        [840] := 2776, [841] := 2780, [842] := 2778, [843] := 2773, [844] := 2778, [845] := 2776, [846] := 2780, [847] := 2783, [848] := 2766, [849] := 2787, [850] := 2773, [851] := 2776, [852] := 2773, [853] := 2780, [854] := 2771, [855] := 2778, [856] := 2771, [857] := 2776, [858] := 2780, [859] := 2785, [860] := 2776, [861] := 2783, [862] := 2776, [863] := 2780, [864] := 2766, [865] := 2776, [866] := 432, [867] := 432, [868] := 2806, [869] := 2797, [870] := 2773, [871] := 531, [872] := 2776, [873] := 2792, [874] := 2790, [875] := 2783, [876] := 2778, [877] := 2780, [878] := 2776, [879] := 2780, [880] := 2771, [881] := 2769, [882] := 2778, [883] := 2780, [884] := 2769, [885] := 2785, [886] := 2776, [887] := 2790, [888] := 2769, [889] := 2785, [890] := 2773, [891] := 2785, [892] := 2776, [893] := 2783, [894] := 2780, [895] := 2785, [896] := 2773, [897] := 2785, [898] := 2778, [899] := 2679,
        [900] := 2691, [901] := 2688, [902] := 2679, [903] := 2676, [904] := 2679, [905] := 2676, [906] := 2679, [907] := 2679, [908] := 2688, [909] := 2691, [910] := 2679, [911] := 2674, [912] := 2681, [913] := 2674, [914] := 2679, [915] := 2681, [916] := 2686, [917] := 2688, [918] := 2693, [919] := 2686, [920] := 2679, [921] := 2674, [922] := 2674, [923] := 2674, [924] := 2743, [925] := 2773, [926] := 2787, [927] := 2776, [928] := 2790, [929] := 2776, [930] := 2776, [931] := 2778, [932] := 2778, [933] := 2771, [934] := 2783, [935] := 2771, [936] := 2780, [937] := 2773, [938] := 2778, [939] := 2769, [940] := 2780, [941] := 2776, [942] := 2776, [943] := 2776, [944] := 2773, [945] := 2785, [946] := 2778, [947] := 2776, [948] := 2776, [949] := 2773, [950] := 2776, [951] := 2778, [952] := 2773, [953] := 2785, [954] := 2771, [955] := 2790, [956] := 2776, [957] := 2764, [958] := 2769, [959] := 2769,
        [960] := 2766, [961] := 2759, [962] := 2761, [963] := 2764, [964] := 2761, [965] := 2776, [966] := 2783, [967] := 2766, [968] := 2757, [969] := 2752, [970] := 2752, [971] := 2754, [972] := 2754, [973] := 2754, [974] := 2750, [975] := 2747, [976] := 2745, [977] := 2754, [978] := 2752, [979] := 2766, [980] := 2761, [981] := 2761, [982] := 2764, [983] := 2764, [984] := 2757, [985] := 2752, [986] := 2766, [987] := 2759, [988] := 2759, [989] := 2771, [990] := 2752, [991] := 2752, [992] := 2752, [993] := 2750, [994] := 2773, [995] := 2771, [996] := 2757, [997] := 2759, [998] := 2754, [999] := 777);
   NEXT_SYNC : ALIAS FOR N7[3];
   O : INT[128] := ([0] := 2#0000_0111_1111_1111, [20] := 2#0000_0010_1000_1000, [21] := 2#0000_0000_0001_0000, [22] := 2#0000_0001_1000_0000, [25] := 2#0000_0000_0001_0000, [26] := 2#0000_0000_0000_0001, [27] := 2#0000_0000_0100_0000, [29] := 2#0000_0000_0001_0000, [33] := 2#0000_0000_0101_0000, [35] := 2#0000_0100_0000_0000, [47] := 2#0000_0100_0000_0000, [59] := 2#0000_0000_0000_0010, [63] := 2#0000_0000_1000_0010, [66] := 2#0010_0000_0000_0000, [67] := 2#0011_1100_0000_0000, [70] := 2#0000_0100_0000_0000, [73] := 2#0000_0000_0000_0001, [78] := 2#0001_0000_0000_0000, [82] := 2#0000_0000_0000_0011, [114] := 2#1001_0010_0100_1001, [115] := 2#1001_0010_0100_0000, [116] := 2#1001_0000_0000_0101, [117] := 2#0000_0000_0001_0000, [118] := 2#1001_0000_0000_0000, [121] := 2#0000_0100_1101_0010, [123] := 2#0000_0000_0001_0010, [124] := 2#0000_1010_0111_1011, [125] := 2#0000_0000_0000_0001);
        [1]   // Scanner 1 Outputs
        [2]   // Scanner 1 Outputs
        [3]   // Scanner 2 Outputs
        [4]   // Scanner 2 Outputs
        [5]   // Scanner 3 Outputs
        [6]   // Scanner 3 Outputs
        [7]   // Scanner 4 Outputs
        [8]   // Scanner 4 Outputs
        [9]   // Scanner 5 Outputs
        [10]   // Scanner 5 Outputs
        [10].15   // Gun 5-11 Shift
        [20].1   // South Chilled Water Blower Start LT I02112 PB
        [20].0   // South Chilled Water Blower Start VFD
        [20].2   // South Chilled Water VFD Stop
        [20].3   // VMCC MB Alarm-horn Relay
        [20].4   // North Chilled Water Blower Start VFD
        [20].5   // North Chilled Water Blower Start LT I02104 PB
        [20].6   // North Chilled Water VFD Stop
        [20].8   // LUCOR MACHINE Operate
        [20].11   // SUB-SURFACE Cutters Raise for Crossbreak Relay
        [20].12   // ISRA 5D System Cut Signal
        [20].13   // ISRA 5D System QC Request Signal
        [21].8   // Temporary Blippy pulse
        [20].14   // Spare
        [20].15   // Spare
        [11].1   // Cullet System Fault Pilot Light (NOT USED ANYMORE)
        [11]   // Lights & Horn (NOT USED ANYMORE)
        [11].0   // Reliance Drive System Fault Pilot Light (NOT USED ANYMORE)
        [25].0   // CRSSBRK ZONE 1 North Outside Lamp
        [25].1   // CRSSBRK ZONE 1 North Inside Lamp
        [25].2   // CRSSBRK ZONE 1 South Outside Lamp
        [25].3   // CRSSBRK ZONE 1 South Inside Lamp
        [25].4   // CRSSBRK ZONE 1 Crossbreak In progress Lamp
        [25].5   // M37B Conv Forward Pilot Light
        [25].6   // M37B Conv Reverse Pilot Light
        [25].7   // M47B Conv Forward Pilot Light
        [25].8   // M47B Conv Reverse Pilot Light
        [27].0   // CRSSBRK ZONE 2 North Outside Lamp
        [27].1   // CRSSBRK ZONE 2 North Inside Lamp
        [27].2   // CRSSBRK ZONE 2 South Outside Lamp (Bad Output)
        [27].3   // CRSSBRK ZONE 2 South Inside Lamp
        [27].4   // CRSSBRK ZONE 2 Crossbreak In progress Lamp
        [27].5   // CRSSBRK ZONE 1 Crossbreak horn Located on wall At lehr Exit
        [27].6   // CRSSBRK ZONE 1 Alarm rotating Beacon Located on lehr Exit
        [27].7   // Crusher #1 Is Lowered (This Output is Read by HE for Pan-alarm Display)
        [27].8   // CRSSBRK ZONE 2 South Outside Lamp (New Output)
        [29].0   // CRSSBRK ZONE 3 North Outside Lamp
        [29].1   // CRSSBRK ZONE 3 North Inside Lamp
        [29].2   // CRSSBRK ZONE 3 South Outside Lamp
        [29].3   // CRSSBRK ZONE 3 South Inside Lamp
        [29].4   // CRSSBRK ZONE 3 Crossbreak In progress Lamp
        [31].6   // IMAGE AUTO Retro cover Manual mode Lamp
        [31].7   // IMAGE AUTO Retro cover Closed Alarm Horn
        [31].8   // IMAGE AUTO Retro cover Alarm Beacon
        [31].10   // IMAGE AUTO Retro Cover Open solenoid Valve
        [33].0   // CRSSBRK ZONE 5 North Outside Lamp
        [33].1   // CRSSBRK ZONE 5 North Inside Lamp
        [33].2   // CRSSBRK ZONE 5 South Outside Lamp
        [33].3   // CRSSBRK ZONE 5 South Inside Lamp
        [33].4   // CRSSBRK ZONE 5 Crossbreak In progress Lamp
        [33].5   // APC Enable Relay
        [33].6   // APC Cut Off relay New Apc Sprayer
        [33].7   // APC #2 Blow off Excess APC During Crossbreak
        [33].8   // APC #2 Lower Roll (On Glass)
        [33].9   // APC #1 Blow off Excess APC During Crossbreak changed 22Mar2019TC
        [33].10   // APC #1 Lower Roll (On Glass) new22MarTC
        [33].11   // APC APC Roll SS1 changed 22Mar2019TC
        [35]   // MANUAL INSPCTN Reject flaw Q.A. flaw Lamps Output word
        [35].0   // MANUAL INSPCTN North Outside Reject Flaw Red Lamp
        [35].1   // MANUAL INSPCTN North Outside Q.A. Flaw Yellow Lamp
        [35].2   // MANUAL INSPCTN North Inside Reject Flaw Red Lamp
        [35].3   // MANUAL INSPCTN North Inside Q.A. Flaw Yellow Lamp
        [35].4   // MANUAL INSPCTN * Center Reject Flaw Red Lamp
        [35].5   // MANUAL INSPCTN * Center Q.A. Flaw Yellow Lamp
        [35].6   // MANUAL INSPCTN South Inside Reject Flaw Red Lamp
        [35].7   // MANUAL INSPCTN South Inside Q.A. Flaw Yellow Lamp
        [35].8   // MANUAL INSPCTN South Outside Reject Flaw Red Lamp
        [35].9   // MANUAL INSPCTN South Outside Q.A. Flaw Yellow Lamp
        [35].10   // MANUAL INSPCTN Cross-break Signal to STP
        [35].11   // MANUAL INSPCTN SPARE
        [35].12   // MANUAL INSPCTN SPARE
        [35].13   // MANUAL INSPCTN * * Function Lamp Clear
        [35].14   // MANUAL INSPCTN * * Function Lamp Blue
        [35].15   // MANUAL INSPCTN Quality Defect Inhibit Function Lamp Red
        [36].0   // RIBBON WASHER AIR KNIFE #2 Converge Solenoid valve NuPlex Block
        [36].2   // RIBBON WASHER AIR KNIFE #1 Converge Solenoid valve NuPlex Block
        [36].4   // RIBBON WASHER SPONGE LOWER Converge Solenoid valve
        [36].6   // RIBBON WASHER SPONGE UPPER Converge Solenoid valve
        [36].8   // RIBBON WASHER TOP HEADER SHUT OFF VALVE
        [36].12   // RIBBON WASHER BRUSH #1 LOWER Converge Solenoid valve
        [36].14   // RIBBON WASHER BRUSH #1 UPPER Converge Solenoid valve
        [45].0   // VMCC W1 Upper Brush #1 Foward
        [45].1   // VMCC W1 Lower Brush #1 Foward
        [45].2   // VMCC W1 Upper Brush #2 Foward
        [47].0   // SPARE
        [45].4   // VMCC W1 Upper Sponge Foward
        [45].5   // VMCC W1 Lower Sponge Foward
        [45].6   // VMCC W1 SPARE
        [45].7   // VMCC W1 SPARE
        [45].8   // VMCC W1 Upper Brush #1 Reverse
        [45].9   // VMCC W1 Lower Brush #1 Reverse
        [45].10   // VMCC W1 Upper Brush #2 Reverse
        [59].10   // SPARE
        [59].1   // SPARE
        [59].5   // SPARE
        [45].14   // VMCC W1 SPARE
        [45].15   // VMCC W1 SPARE
        [46].0   // VMCC W1 Upper Brush #1 Speed Select 1
        [63].13   // SPARE
        [46].2   // VMCC W1 Upper Brush #2 Speed Select 1
        [63].12   // SPARE
        [59].7   // PANEL W2 AIR KNIFE RELAY AKBR-ON
        [63].14   // SPARE
        [46].6   // VMCC W1 SPARE
        [46].7   // VMCC W1 SPARE
        [46].8   // VMCC W1 Upper Brush #1 Speed Select 2
        [46].9   // VMCC W1 Lower Brush #1 Speed Select 2
        [46].10   // VMCC W1 Upper Brush #2 Speed Select 2
        [63].11   // SPARE
        [46].13   // VMCC W1 Lower Sponge Speed Select 2
        [46].14   // VMCC W1 SPARE
        [46].15   // VMCC W1 SPARE
        [47].13   // SPARE
        [59].8   // SPARE
        [47].11   // SPARE
        [47].12   // SPARE
        [47].14   // SPARE
        [47].4   // VMCC W1 Blue Stack Light (NOT USED ANYMORE)
        [47].15   // SPARE
        [47].8   // VMCC W1 Water Sprayer #2 ON (This is the spray bar)
        [47].9   // VMCC W1 Water Sprayer #3 ON
        [47].10   // CRSSBRK ZONE 1 Alarm Rotating Beacon Located In Acid Washer Room
        [59].0   // PANEL W2 BRUSH #1 Manual mode Lamp
        [59].2   // PANEL W2 SPONGE UNIT Manual mode Lamp
        [59].3   // PANEL W2 AIR KNIVES Manual mode Lamp
        [59].4   // PANEL W2 WATER SPRAYERS Manual mode Lamp
        [63].5   // SPARE
        [63].1   // SPARE
        [63].0   // PANEL W3 BRUSH #1 Manual mode Lamp
        [63].2   // PANEL W3 SPONGE UNIT Manual mode Lamp
        [63].3   // PANEL W3 AIR KNIVES Manual mode Lamp
        [63].4   // PANEL W3 WATER SPRAYERS Manual mode Lamp
        [63].15   // SPARE
        [66].0   // VMCC M1 Crusher #1 Forward
        [66].2   // VMCC M1 Crusher #1 Speed Select 1
        [66].4   // VMCC M1 Crusher #1 Speed Select 2
        [66].6   // VMCC M1 Crusher #1 Speed Select 3
        [66].8   // VMCC M1 Drive Fault Lamp
        [66].9   // VMCC M1 Drive Fault Reset relay
        [66].13   // VMCC M1 Alarm Horn Relay
        [67].0   // VMCC M1 Crusher #1 Up Relay
        [67].1   // VMCC M1 Crusher #1 Down Relay
        [67].3   // VMCC M1 Red Stack Lite
        [67].4   // VMCC M1 Blue Stack Lite
        [67].5   // VMCC M1 Amber Stack Lite
        [67].8   // VMCC M1 Crusher #1 ON Lamp
        [67].9   // VMCC M1 Crusher #1 OFF Lamp
        [67].10   // BAD OUTPUT 12 TERMINAL 10- DO NOT USE
        [67].11   // No. 1 Crusher Chip Blower On Pilot Light (Top)
        [67].12   // No. 1 Crusher Chip Blower On Pilot Light (VMCC M1)
        [67].13   // No. 1 Crusher Chip Blower 24VDC Relay for M1 Coil
        [82].0   // RELIANCE DRIVE PANEL Permissive to Run from PLC MB
        [82].1   // RELIANCE DRIVE PANEL Permissive to Run from PLC MB Stops on line/bk
        [112].12   // MB --> Cullet Diverter Position at Bin 1B
        [113].14   // CULLET SYSTEM VP 917067 Vibrating pan Thin glass Speed
        [113].15   // CULLET SYSTEM VP 917067 Vibrating pan Medium glass Speed
        [114].0   // CULLET SYSTEM VP 917067 Vibrating pan Thick glass Speed
        [114].1   // CULLET SYSTEM VP 917066 Vibrating pan Thin glass Speed
        [114].2   // CULLET SYSTEM VP 917066 Vibrating pan Medium glass Speed
        [114].3   // CULLET SYSTEM VP 917066 Vibrating pan Thick glass Speed
        [114].4   // CULLET SYSTEM VP 917065 Vibrating pan Thin glass Speed
        [114].5   // CULLET SYSTEM VP 917065 Vibrating pan Medium glass Speed
        [114].6   // CULLET SYSTEM VP 917065 Vibrating pan Thick glass Speed
        [114].7   // CULLET SYSTEM VP 917070 Vibrating pan Thin glass Speed
        [114].8   // CULLET SYSTEM VP 917070 Vibrating pan Medium glass Speed
        [114].9   // CULLET SYSTEM VP 917070 Vibrating pan Thick glass Speed
        [114].10   // CULLET SYSTEM VP 917071 Vibrating pan Thin glass Speed
        [114].11   // CULLET SYSTEM VP 917071 Vibrating pan Medium glass Speed
        [114].12   // CULLET SYSTEM VP 917071 Vibrating pan Thick glass Speed
        [114].13   // CULLET SYSTEM VP 917077 Vibrating pan Thin glass Speed
        [114].14   // CULLET SYSTEM VP 917077 Vibrating pan Medium glass Speed
        [114].15   // CULLET SYSTEM VP 917077 Vibrating pan Thick glass Speed
        [115].1   // MB --> Cullet ML is in Sleep Mode
        [115].2   // MB --> Cullet Leg 4 Is In Sleep Mode
        [118].14   // MB --> Cullet ???
        [115].4   // CULLET SYSTEM VP 917076 Vibrating pan Thin glass Speed
        [115].5   // CULLET SYSTEM VP 917076 Vibrating pan Medium glass Speed
        [115].6   // CULLET SYSTEM VP 917076 Vibrating pan Thick glass Speed
        [115].7   // CULLET SYSTEM VP 917075 Vibrating pan Thin glass Speed
        [115].8   // CULLET SYSTEM VP 917075 Vibrating pan Medium glass Speed
        [115].9   // CULLET SYSTEM VP 917075 Vibrating pan Thick glass Speed
        [115].10   // CULLET SYSTEM VP 917074 Vibrating pan Thin glass Speed
        [115].11   // CULLET SYSTEM VP 917074 Vibrating pan Medium glass Speed
        [115].12   // CULLET SYSTEM VP 917074 Vibrating pan Thick glass Speed
        [115].13   // CULLET SYSTEM VP 917073 Vibrating pan Thin glass Speed
        [115].14   // CULLET SYSTEM VP 917073 Vibrating pan Medium glass Speed
        [115].15   // CULLET SYSTEM VP 917073 Vibrating pan Thick glass Speed
        [116].2   // CULLET SYSTEM VP 917069 Vibrating pan Thick glass Spee
        [116].7   // CULLET SYSTEM VP 917068 Vibrating pan Thick glass Speed
        [116].8   // CULLET SYSTEM Diverter Position 1
        [116].10   // CULLET SYSTEM VP 917072 Vibrating pan Thin glass Speed
        [116].11   // CULLET SYSTEM VP 917072 Vibrating pan Medium glass Speed
        [116].12   // CULLET SYSTEM VP 917072 Vibrating pan Thick glass Speed
        [116].13   // CULLET SYSTEM VP 917060 Vibrating pan Thin glass Speed
        [116].14   // CULLET SYSTEM VP 917060 Vibrating pan Medium glass Speed
        [116].15   // CULLET SYSTEM VP 917060 Vibrating pan Thick Glass Speed crusher #1 VP
        [119].4   // MB --> C1 Float Glass Production
        [117].15   // MB --> Cullet PANEL C3 M-41 CONVEYOR SLEEP MODE
        [118].1   // MB --> Cullet Leg 3 Is In Sleep Mode Turn Off Belt 3 of 3
        [118].10   // MB --> Cullet Crusher No. 2 Is Operating
        [118].12   // MB --> Cullet Crusher No. 3 Is Operating
        [119].0   // MB --> Cullet M37B Run Fwd Signal
        [119].1   // MB --> Cullet M37B Run Rev Signal
        [119].2   // MB --> Cullet M47B Run Fwd Signal
        [119].3   // MB --> Cullet M47B Run Rev Signal
        [119].5   // From Host Enable 37B's REV controls
        [123].1   // MB -->> M2 Crossbreak In progress Front end
        [123].3   // MB -->> M2 No. 1 Crusher Down prox. Made
        [123].4   // MB -->> M2 Eclipse Mode Signal For Hold Down Wheels
        [123].5   // MB -->> M2 Sub-surface Cutters In Alarm
        [125]   // MB -->> M2 Host comp. Reliance Crossbreaks Disable Ycuts
        [125].0   // MB -->> M2 Crossbreak Signal to Reliance Capping system
        [31].0   // CRSSBRK ZONE 4 North Outside Lamp
        [20].9   // Spare
        [59].13   // SPARE
        [59].11   // SPARE
        [59].12   // SPARE
        [63].10   // SPARE
        [59].14   // SPARE
        [47].1   // VMCC W1 Drive fault Lamp (NOT USED ANYMORE)
        [47].5   // VMCC W1 Amber Stack Light (NOT USED ANYMORE)
        [63].9   // SPARE
        [63].7   // SPARE
        [59].9   // SPARE
        [59].15   // SPARE
        [47].7   // VMCC W1 Water Sprayer #1 ON (NOT USED ANYMORE)
        [63].6   // PANEL W3 AIR KNIFE SS LIGHT ON PANEL #W3
        [47].3   // VMCC W1 Red Stack Light (NOT USED ANYMORE)
        [59].6   // PANEL W2 AIR KNIFE SS LIGHT ON PANEL #W2
        [63].8   // SPARE
        [33]   // CRSSBRK ZONE 5 & APC
        [118].15   // MB --> Cullet ???
        [20]   // Water SUB-SURFACE ISRA
        [63]   // PANEL W3
        [66]   // VMCC M1
        [67]   // VMCC M1
        [123]   // MB --> M2
        [124]   // MB --> M2
        [82]   // RELIANCE DRIVE PANEL
        [29]   // CRSSBRK ZONE 3
        [31]   // IMAGE AUTO
        [36]   // RIBBON WASHER
        [112]   // MB --> Cullet
        [31].1   // CRSSBRK ZONE 4 North Inside Lamp
        [31].2   // CRSSBRK ZONE 4 South Outside Lamp
        [31].3   // CRSSBRK ZONE 4 South Inside Lamp
        [31].4   // CRSSBRK ZONE 4 Crossbreak In progress Lamp
        [31].9   // IMAGE AUTO Open Graticule Solenoid (Raise)
        [45]   // VMCC W1
        [118]   // MB --> Cullet
        [113]   // MB --> Cullet
        [46]   // VMCC W1
        [47]   // VMCC W1
        [20].10   // Spare
        [119]   // MB --> Cullet
        [25]   // CRSSBRK ZONE 1
        [114]   // MB --> Cullet
        [115]   // MB --> Cullet
        [27]   // CRSSBRK ZONE 2
        [116]   // MB --> Cullet
        [20].7   // Spare
        [59]   // PANEL W2
        [117]   // MB --> Cullet
        [22]   // Lamps (NOT USED ANYMORE)
        [22].3   // MARKING BRIDGE Lower Lamp (NOT USED ANYMORE)
        [22].4   // Bridge in Spray Position Lamp (NOT USED ANYMORE)
        [22].7   // CRSSBRK ZONE 5 APC (MAN INSPECT) Crossbreak In progress Lamp at Capping (NOT USED ANYMORE)
        [22].8   // CRSSBRK ZONE 1 Lehr Crossbreak In progress Lamp at Capping (NOT USED ANYMORE)
        [22].9   // CRSSBRK ZONE 2 Lehr exit Crossbreak In progress Lamp at Capping (NOT USED ANYMORE)
        [11].2   // Reliance Drive & Cullet System Alarm Horn Relay (Capping Rm) (NOT USED ANYMORE)
        [45].3   // VMCC W1 Lower Brush #2 Foward (NOT USED ANYMORE)
        [45].12   // VMCC W1 Upper Sponge Reverse (NOT USED ANYMORE)
        [45].11   // VMCC W1 Lower Brush #2 Reverse (NOT USED ANYMORE)
        [45].13   // VMCC W1 Lower Sponge Reverse (NOT USED ANYMORE)
        [46].1   // VMCC W1 Lower Brush #1 Speed Select 1 (NOT USED ANYMORE)
        [46].3   // VMCC W1 Lower Brush #2 Speed Select 1 (NOT USED ANYMORE)
        [46].4   // VMCC W1 Upper Sponge Speed Select 1 (NOT USED ANYMORE)
        [46].5   // VMCC W1 Lower Sponge Speed Select 1 (NOT USED ANYMORE)
        [46].11   // VMCC W1 Lower Brush #2 Speed Select 2 (NOT USED ANYMORE)
        [46].12   // VMCC W1 Upper Sponge Speed Select 2
        [47].2   // VMCC W1 Drive fault Reset relay
        [47].6   // VMCC W1 Mainline ??? Matt Tipping What is it?
        [115].0   // MB --> Cullet PANEL C4 M34t MAIN #1 CONV SLEEP MODE
        [115].3   // MB --> Cullet PANEL C4 M-33 CONVEYOR SLEEP MODE; TURN OFF LEG #5
        [117].4   // MB --> Cullet #1 CRUSHER RUNNING; ENABLE VP 917060 FOR DISCHARGE
        [117].14   // MB --> Cullet PANEL C3 M-43 CONVEYOR SLEEP MODE; TURN OFF LEG #2
        [118].0   // MB --> Cullet PANEL C3 M-42 CONVEYOR SLEEP MODE; TURN OFF LEG #3
        [118].13   // MB --> Cullet #4 CRUSHER RUNNING; ENABLE VP 917068 TO RUN
   ProducedToCullet : UDT_PRODUCED_CULLET := (MBtoCULLET_3 := -28087, MBtoCULLET_4 := -28096, MBtoCULLET_5 := -28667, MBtoCULLET_6 := 16, MBtoCULLET_7 := -28672);
   ProducedToMCC1300 : UDT_PRODUCED_NEXT := (iMBtoM2_2 := 1234, iMBtoM2_4 := 18, iMBtoM2_5 := 2683, iMBtoM2_6 := 1); {produced}
   R150 : CONTROL[6] := ([1].LEN := 48, [1].UL := 1, [2].LEN := 600, [3].LEN := 72, [3].UL := 1, [4].LEN := 148, [5].LEN := 240, [5].UL := 1);
        [1]   // Control for Cross-break Zone 1 Bit shift Tracking
        [2]   // Control for Cross-break Zone 2 Bit shift Tracking
        [3]   // Control for Cross-break Zone 3 Bit shift Tracking
        [4]   // Control for Cross-break Zone 4 Bit shift Tracking
        [5]   // Control for Cross-break Zone 5 Bit shift Tracking
   R509 : CONTROL[2] := ([0].LEN := 7, [1].LEN := 2, [1].POS := 1, [1].EN := 1, [1].DN := 1);
        [1]   // SPEED CALC FAL control For washer Sponge Drives
   R509_000_POS : ALIAS FOR R509[0].POS;
   R509_001_POS : ALIAS FOR R509[1].POS;
   R56 : CONTROL[20];
   R6 : CONTROL[100] := ([0].LEN := 1000, [0].POS := 999, [0].EN := 1, [0].DN := 1);
   R97 : CONTROL[4] := ([0].LEN := 10, [1].LEN := 10);
        [0]   // LEHR SPEED Control word For Lehr Speed averaging Function
        [1]   // LEHR SPEED Control word For lehr Speed standard Deviation
   REG_INDEX : DINT := 382; {access Read Only}
   REL_2IN_PULSE : ALIAS FOR N54[301].1;
   REL_CAP_REQUEST : ALIAS FOR I[17].14;
   REL_DATA_REQ : ALIAS FOR N54[301].0;
   REL_DRV_FLT : ALIAS FOR B3[3].0;
   RELDR_ESTOP : ALIAS FOR I[80].0;
   RELIANCE_FLT_PL : ALIAS FOR O[11].0;
   S : INT[128] := ([0] := 16#0004, [1] := 16#2082, [2] := 16#ca4c, [7] := 16#0008, [8] := 16#0016, [9] := 16#0035, [10] := 16#5004, [13] := 16#0002, [14] := 16#002d, [16] := 16#00bc, [17] := 16#0200, [18] := 16#07e7, [19] := 16#0006, [20] := 16#0009, [21] := 16#000f, [22] := 16#0011, [23] := 16#0005, [28] := 16#01f4, [30] := 16#000a, [31] := 16#0012, [46] := 16#0013, [47] := 16#000d, [48] := 16#0001, [49] := 16#0001, [51] := 16#0001, [53] := 16#0001, [54] := 16#0005, [55] := 16#0001, [56] := 16#0002, [57] := 16#7a3b, [64] := 16#0003, [76] := 16#0004, [78] := 16#fbe7, [79] := 16#3064, [80] := 16#0002, [81] := 16#000a, [82] := 16#001e, [83] := 16#0003, [85] := 16#000d, [88] := 16#0011, [94] := 16#000e, [95] := 16#0007, [97] := 16#0013, [98] := 16#0008, [101] := 16#0009, [102] := 16#0002, [103] := 16#000b, [104] := 16#000a, [105] := 16#0001, [106] := 16#0008, [107] := 16#000b, [108] := 16#0003, [109] := 16#0007, [110] := 16#000c, [111] := 16#0002, [112] := 16#000c, [113] := 16#000d, [114] := 16#0003, [115] := 16#0014, [116] := 16#000e,
        [119] := 16#000f, [122] := 16#0010, [123] := 16#0001, [124] := 16#0007, [125] := 16#0011, [126] := 16#0005, [127] := 16#0013);
        [0].0   // Processor arithmetic carry flag
        [0].1   // Processor arithmetic underflow/ overflow flag
        [0].2   // Processor arithmetic zero flag
        [0].3   // Processor arithmetic sign flag
        [1].0   // Bad RAM CHECKSUM at power up
        [1].1   // PLC-5 in RUN mode
        [1].2   // PLC-5 in TEST mode
        [1].3   // PLC-5 in PROG mode
        [1].4   // PLC-5 is burning an EEPROM
        [1].5   // Download- ing in progress
        [1].6   // Test edits enabled
        [1].7   // Mode switch in REMOTE
        [1].8   // Forces enabled
        [1].9   // Forces present
        [1].10   // EEPROM success- fully Burned
        [1].11   // Perform- ing online program- ming
        [1].12   // Processor is in DEBUG mode
        [1].13   // User program CHECKSUM done
        [1].14   // Last scan of ladder or SFC step
        [1].15   // First Scan
        [7].0   // Rack 0 Faulted
        [7].1   // Rack 1 Faulted
        [7].2   // Rack 2 Faulted
        [7].3   // Rack 3 Faulted
        [7].4   // Rack 4 Faulted
        [7].5   // Rack 5 Faulted
        [7].6   // Rack 6 Faulted
        [7].7   // Rack 7 Faulted
        [7].8   // Block Xfer queue to rack 0 is full
        [7].9   // Block Xfer queue to rack 1 is full
        [7].10   // Block Xfer queue to rack 2 is full
        [7].11   // Block Xfer queue to rack 3 is full
        [7].12   // Block Xfer queue to rack 4 is full
        [7].13   // Block Xfer queue to rack 5 is full
        [7].14   // Block Xfer queue to rack 6 is full
        [7].15   // Block Xfer queue to rack 7 is full
        [8]   // Last program scan time ladder & SFC
        [9]   // Maximum program scan time ladder & SFC
        [10].0   // Battery is bad or missing
        [10].1   // DH+ active node table changed
        [10].2   // STI overlap
        [10].3   // EEPROM trans- ferred
        [10].4   // Edits prevent SFC continuing
        [10].5   // Invalid I/O status file
        [10].6   // Memory cartridge battery low
        [10].7   // No more command blocks exist
        [10].9   // No MCP was configured to run
        [10].10   // MCP not allowed
        [10].11   // PII word number isn't in local rack
        [10].12   // User PII routine overlap
        [10].13   // No command block exists to get PII
        [10].14   // Arithmetic overflow occurred
        [10].15   // SFC lingering action overlap
        [11].0   // Bad program file
        [11].1   // Bad address in ladder program
        [11].2   // Programmer error
        [11].3   // SFC Fault
        [11].4   // Program assembly error
        [11].5   // Powerup protection fault
        [11].6   // Error not defined
        [11].7   // User generated fault
        [11].8   // Watchdog timer fault
        [11].9   // Bad system config- uration
        [11].10   // Hardware Error
        [11].11   // MCP file does not exist or is not ladder
        [11].12   // PII file does not exist or is not ladder
        [11].13   // STI file does not exist or is not ladder
        [11].14   // Fault file does not exist or is not ladder
        [11].15   // Non ladder file
        [12]   // Fault Code
        [13]   // Program file where fault occurred
        [14]   // Rung number where fault occurred
        [16]   // I/O status file
        [17].0   // Queue full between local and remote I/O
        [17].1   // Queue full servicing channel 1A
        [17].2   // Queue full servicing channel 1B
        [17].3   // Queue full servicing channel 2A
        [17].4   // Queue full servicing channel 2B
        [17].5   // No modem on serial port
        [17].6   // Remote I/O is greater than image size
        [17].8   // ASCII instruct- ion error
        [17].9   // Duplicate node address
        [18]   // Real time clock YEAR
        [19]   // Real time clock MONTH
        [20]   // Real time clock DAY
        [21]   // Real time clock HOUR
        [22]   // Real time clock MINUTE
        [23]   // Real time clock SECOND
        [24]   // Index Offset
        [25]   // Adapter Image File
        [26].0   // SFC Restart/ Continue
        [26].1   // Start-up protect- ion after power loss
        [26].2   // Local rack is 1 if set or 0 if bit = 0
        [26].3   // Complement Rack Mode
        [27].0   // Rack 0 Inhibit
        [27].1   // Rack 1 Inhibit
        [27].2   // Rack 2 Inhibit
        [27].3   // Rack 3 Inhibit
        [27].4   // Rack 4 Inhibit
        [27].5   // Rack 5 Inhibit
        [27].6   // Rack 6 Inhibit
        [27].7   // Rack 7 Inhibit
        [27].8   // Rack 0 Reset
        [27].9   // Rack 1 Reset
        [27].10   // Rack 2 Reset
        [27].11   // Rack 3 Reset
        [27].12   // Rack 4 Reset
        [27].13   // Rack 5 Reset
        [27].14   // Rack 6 Reset
        [27].15   // Rack 7 Reset
        [28]   // Watchdog Timer Setpoint
        [29]   // Fault routine file number
        [30]   // STI setpoint (interval)
        [31]   // STI file number
        [32].0   // Rack 10 Faulted
        [32].1   // Rack 11 Faulted
        [32].2   // Rack 12 Faulted
        [32].3   // Rack 13 Faulted
        [32].4   // Rack 14 Faulted
        [32].5   // Rack 15 Faulted
        [32].6   // Rack 16 Faulted
        [32].7   // Rack 17 Faulted
        [32].8   // Block Xfer queue to rack 10 is full
        [32].9   // Block Xfer queue to rack 11 is full
        [32].10   // Block Xfer queue to rack 12 is full
        [32].11   // Block Xfer queue to rack 13 is full
        [32].12   // Block Xfer queue to rack 14 is full
        [32].13   // Block Xfer queue to rack 15 is full
        [32].14   // Block Xfer queue to rack 16 is full
        [32].15   // Block Xfer queue to rack 17 is full
        [33].0   // Rack 10 Inhibit
        [33].1   // Rack 11 Inhibit
        [33].2   // Rack 12 Inhibit
        [33].3   // Rack 13 Inhibit
        [33].4   // Rack 14 Inhibit
        [33].5   // Rack 15 Inhibit
        [33].6   // Rack 16 Inhibit
        [33].7   // Rack 17 Inhibit
        [33].8   // Rack 10 Reset
        [33].9   // Rack 11 Reset
        [33].10   // Rack 12 Reset
        [33].11   // Rack 13 Reset
        [33].12   // Rack 14 Reset
        [33].13   // Rack 15 Reset
        [33].14   // Rack 16 Reset
        [33].15   // Rack 17 Reset
        [34].0   // Rack 20 Faulted
        [34].1   // Rack 21 Faulted
        [34].2   // Rack 22 Faulted
        [34].3   // Rack 23 Faulted
        [34].4   // Rack 24 Faulted
        [34].5   // Rack 25 Faulted
        [34].6   // Rack 26 Faulted
        [34].7   // Rack 27 Faulted
        [34].8   // Block Xfer queue to rack 20 is full
        [34].9   // Block Xfer queue to rack 21 is full
        [34].10   // Block Xfer queue to rack 22 is full
        [34].11   // Block Xfer queue to rack 23 is full
        [34].12   // Block Xfer queue to rack 24 is full
        [34].13   // Block Xfer queue to rack 25 is full
        [34].14   // Block Xfer queue to rack 26 is full
        [34].15   // Block Xfer queue to rack 27 is full
        [35].0   // Rack 20 Inhibit
        [35].1   // Rack 21 Inhibit
        [35].2   // Rack 22 Inhibit
        [35].3   // Rack 23 Inhibit
        [35].4   // Rack 24 Inhibit
        [35].5   // Rack 25 Inhibit
        [35].6   // Rack 26 Inhibit
        [35].7   // Rack 27 Inhibit
        [35].8   // Rack 20 Reset
        [35].9   // Rack 21 Reset
        [35].10   // Rack 22 Reset
        [35].11   // Rack 23 Reset
        [35].12   // Rack 24 Reset
        [35].13   // Rack 25 Reset
        [35].14   // Rack 26 Reset
        [35].15   // Rack 27 Reset
        [46]   // PII file number
        [47]   // PII module group to examine
        [48]   // PII bit mask
        [48].0   // PII Module Bit 1=Monitor 0=Ignore
        [49]   // PII compare value
        [49].0   // PII Bit 1=false to TRUE 0= true to
        [50]   // PII down count
        [51]   // PII return mask
        [52]   // PII accum- ulator
        [53]   // STI last scan time
        [54]   // STI max scan time
        [55]   // PII last scan time
        [56]   // PII max scan time
        [79].0   // Main control program A disable bit
        [79].1   // Main control program B disable bit
        [79].2   // Main control program C disable bit
        [79].3   // Main control program D disable bit
        [79].4   // Main control program E disable bit
        [79].5   // Main control program F disable bit
        [79].6   // Main control program G disable bit
        [79].7   // Main control program H disable bit
        [79].8   // Main control program I disable bit
        [79].9   // Main control program J disable bit
        [79].10   // Main control program K disable bit
        [79].11   // Main control program L disable bit
        [79].12   // Main control program M disable bit
        [79].13   // Main control program N disable bit
        [79].14   // Main control program O disable bit
        [79].15   // Main control program P disable bit
        [80]   // Main control program A file number
        [81]   // Program A scan time
        [82]   // Program A maximum scan time
        [83]   // Main control program B file number
        [84]   // Program B scan time
        [85]   // Program B maximum scan time
        [86]   // Main control program C file number
        [87]   // Program C scan time
        [88]   // Program C maximum scan time
        [89]   // Main control program D file number
        [90]   // Program D scan time
        [91]   // Program D maximum scan time
        [92]   // Main control program E file number
        [93]   // Program E scan time
        [94]   // Program E maximum scan time
        [95]   // Main control program F file number
        [96]   // Program F scan time
        [97]   // Program F maximum scan time
        [98]   // Main control program G file number
        [99]   // Program G scan time
        [100]   // Program G maximum scan time
        [101]   // Main control program H file number
        [102]   // Program H scan time
        [103]   // Program H maximum scan time
        [104]   // Main control program I file number
        [105]   // Program I scan time
        [106]   // Program I maximum scan time
        [107]   // Main control program J file number
        [108]   // Program J scan time
        [109]   // Program J maximum scan time
        [110]   // Main control program K file number
        [111]   // Program K scan time
        [112]   // Program K maximum scan time
        [113]   // Main control program L file number
        [114]   // Program L scan time
        [115]   // Program L maximum scan time
        [116]   // Main control program M file number
        [117]   // Program M scan time
        [118]   // Program M maximum scan time
        [119]   // Main control program N file number
        [120]   // Program N scan time
        [121]   // Program N maximum scan time
        [122]   // Main control program O file number
        [123]   // Program O scan time
        [124]   // Program O maximum scan time
        [125]   // Main control program P file number
        [126]   // Program P scan time
        [127]   // Program P maximum scan time
   Sbr_IN_dDataLength : DINT := 501;
   SFLASH_SLAVE : ALIAS FOR T51[1];
   SLOW_FLASH : ALIAS FOR T51[0];
   SPNGE_DN_FLT : ALIAS FOR I[43].5;
   SPNGE_DN_FWD : ALIAS FOR O[45].5;
   SPNGE_DN_REV : ALIAS FOR O[45].13;
   SPNGE_DN_SS1 : ALIAS FOR O[46].5;
   SPNGE_DN_SS2 : ALIAS FOR O[46].13;
   SPNGE_UP_FLT : ALIAS FOR I[43].4;
   SPNGE_UP_FWD : ALIAS FOR O[45].4;
   SPNGE_UP_REV : ALIAS FOR O[45].12;
   SPNGE_UP_SS1 : ALIAS FOR O[46].4;
   SPNGE_UP_SS2 : ALIAS FOR O[46].12;
   SPRAY_LENGTH : ALIAS FOR N7[8];
   SPRAY_POS_LAMP : ALIAS FOR O[22].4;
   SSW_CAW_OFF_W2 : ALIAS FOR I[58].6;
   SSW_CAW_OFF_W3 : ALIAS FOR I[62].6;
   SSW_CAW_ON_W2 : ALIAS FOR I[58].5;
   SSW_CAW_ON_W3 : ALIAS FOR I[62].5;
   Status : INT := 12384;   // INT tag to retrieve Status value through GSV created during conversion
   STRAIN_CNT : ALIAS FOR N46[0];
   STRAIN_CYC : ALIAS FOR N46[2];
   STRAIN_STAT : ALIAS FOR N46[1];
   T160 : TIMER[100] := ([0].PRE := 100, [0].ACC := 100, [0].EN := 1, [0].DN := 1, [1].PRE := 100, [1].ACC := 100, [1].EN := 1, [1].DN := 1, [2].PRE := 100, [2].ACC := 100, [2].EN := 1, [2].DN := 1, [3].PRE := 100, [3].ACC := 100, [3].EN := 1, [3].DN := 1);
        [0]   // CRSSBRK ZONE 5 North Outside Photo-cell OFF Debounce Timer
        [1]   // CRSSBRK ZONE 5 North Inside Photo-cell OFF Debounce Timer
        [2]   // CRSSBRK ZONE 5 South Outside Photo-cell OFF Debounce Timer
        [3]   // CRSSBRK ZONE 5 South Inside Photo-cell OFF Debounce Timer
   T182 : TIMER[11] := ([0].PRE := 5000, [0].ACC := 5000, [0].EN := 1, [0].DN := 1, [1].PRE := 500, [2].PRE := 10, [3].PRE := 30000, [4].PRE := 10000, [5].PRE := 20000000, [6].PRE := 1000, [9].PRE := 10000, [10].PRE := 100);
   T252 : TIMER[49];
   T4 : TIMER[100] := ([0].PRE := 2500, [1].PRE := 3000, [1].ACC := 3000, [2].PRE := 300, [2].EN := 1, [2].DN := 1, [3].PRE := 327670, [3].ACC := 327670, [3].EN := 1, [3].DN := 1, [4].PRE := 327670, [4].ACC := 327670, [4].EN := 1, [4].DN := 1, [5].PRE := 60000, [5].ACC := 60000, [5].EN := 1, [5].DN := 1, [6].PRE := 15000, [7].PRE := 3000, [7].ACC := 3000, [8].PRE := 2000, [10].PRE := 30000, [11].PRE := 4140, [12].PRE := 4140, [13].PRE := 30000, [17].PRE := 300, [17].ACC := 300, [17].EN := 1, [17].DN := 1, [18].PRE := 200, [18].ACC := 200, [18].EN := 1, [18].DN := 1, [19].PRE := 200, [19].ACC := 200, [19].EN := 1, [19].DN := 1, [20].PRE := 200, [20].ACC := 200, [20].EN := 1, [20].DN := 1, [21].PRE := 200, [21].ACC := 200, [21].EN := 1, [21].DN := 1, [22].PRE := 200, [22].ACC := 200, [22].EN := 1, [22].DN := 1, [23].PRE := 200, [23].ACC := 200, [23].EN := 1, [23].DN := 1, [24].PRE := 250, [24].ACC := 250, [24].EN := 1, [24].DN := 1, [28].PRE := 10, [29].PRE := 20,
        [30].PRE := 20, [31].PRE := 20, [32].PRE := 20, [33].PRE := 500, [33].ACC := 500, [33].EN := 1, [33].DN := 1, [34].PRE := 500, [34].ACC := 500, [34].EN := 1, [34].DN := 1, [35].PRE := 500, [35].ACC := 500, [35].EN := 1, [35].DN := 1, [36].PRE := 350, [36].ACC := 350, [36].EN := 1, [36].DN := 1, [50].PRE := 1500, [50].ACC := 2501, [50].EN := 1, [50].DN := 1, [51].PRE := 1500, [80].PRE := 10, [95].PRE := 500, [96].PRE := 1000, [97].PRE := 500, [98].PRE := 200, [98].ACC := 201, [98].EN := 1, [98].DN := 1, [99].PRE := 4600, [99].ACC := 4601, [99].EN := 1, [99].DN := 1);
        [0]   // Init Timer
        [0].TT   // Initialize
        [1]   // ISRA 5D Off Delay for Error 1
        [2].ACC   // Time of Current Read
        [3]   // Host New Data Timer
        [3].ACC   // Elapsed Time of Current Data
        [4]   // Time Accumulated Since last 1 Meter Pulse
        [4].ACC   // Time accumulate d since last 1 Meter pulse
        [5]   // NO1 CRUSHER Crusher is up and in manual timer.
        [6]   // Capping Room Alarm Horn Relay Duration
        [7]   // ISRA 5D Off Delay for Error 2
        [10]   // South Chilled Water Blower VFD Delay to Restart
        [11]   // TEMP DEBUG OF 1 M SYNC PULSE ON STATE
        [12]   // TEMP DEBUG OF 1 M SYNC PULSE OFF STATE
        [13]   // North Chilled Water Blower VFD Delay to Restart
        [17]   // CRSSBRK ZONE 1 North Outside Photo-cell Off Debounce Timer
        [18]   // CRSSBRK ZONE 1 North Inside Photo-cell Off Debounce Timer
        [19]   // CRSSBRK ZONE 1 South Outside Photo-cell Off Debounce Timer
        [20]   // CRSSBRK ZONE 1 South Inside Photo-cell Off Debounce Timer
        [21]   // CRSSBRK ZONE 2 North Outside Photo-cell Off Debounce Timer
        [22]   // CRSSBRK ZONE 2 North Inside Photo-cell Off Debounce Timer
        [23]   // CRSSBRK ZONE 2 South Outside Photo-cell Off Debounce Timer
        [24]   // CRSSBRK ZONE 2 South Inside Photo-cell Off Debounce Timer
        [28]   // ISRA 5D System Cut Signal Delay
        [33]   // CRSSBRK ZONE 3 North Outside Photo-cell Off Debounce Timer
        [34]   // CRSSBRK ZONE 3 North Inside Photo-cell Off Debounce Timer
        [35]   // CRSSBRK ZONE 3 South Outside Photo-cell Off Debounce Timer
        [36]   // CRSSBRK ZONE 3 South Inside Photo-cell Off Debounce Timer
        [50]   // APC #1 Timer to Blow off excess APC during Crossbreak
        [51]   // APC #2 Timer to Blow off excess APC during Crossbreak
        [95]   // APC #2 Lower Roll Delay Timer
        [96]   // VISION SYS Rejected Plate Alarm Horn
        [97]   // APC #1 Lower Roll Delay Timer
        [98]   // APC #1 Turn on APC Flood Valve Delay
        [99]   // APC #1 Flood Valve Run Time
   T51 : TIMER[13] := ([0].PRE := 750, [0].ACC := 370, [0].EN := 1, [0].TT := 1, [1].PRE := 1000, [2].PRE := 150, [3].PRE := 40, [3].ACC := 20, [3].EN := 1, [3].TT := 1, [9].PRE := 300000, [10].PRE := 50, [10].ACC := 50, [11].PRE := 5000, [12].PRE := 2500, [12].ACC := 2500, [12].EN := 1, [12].DN := 1);
        [0]   // SLOW FLASH Use this timer .EN bit to create slowly flashing lamps
        [0].DN   // SLOW FLASH Use this DoNe bit to create slowly flashing lamps
        [1]   // SLOW FLASH This the slave timer for the slow flash timer
        [2]   // FAST FLASH Use this timer .DN bit to create fast flashing lamps
        [2].DN   // FAST FLASH Use this timer .DoNe bit to create fast flashing lamps
        [2].EN   // FAST FLASH Enable bit for the fast flash timer
        [3]   // FAST FLASH This is the slave timer for the fast flash timer
        [3].DN   // FAST FLASH DoNe bit for fast flash slave timer
        [3].EN   // FAST FLASH Enable bit for the fast flash slave timer
        [9]   // No. 1 Crusher Chip Blower Duration for Automatic Mode
        [11]   // NO. 1 CRUSHER First scan Latch Timer
   T57 : TIMER[100] := ([1].PRE := 100, [2].PRE := 100, [6].PRE := 30000, [6].ACC := 30000, [6].EN := 1, [6].DN := 1, [10].PRE := 300);
        [1]   // Ribbon Washer Brush #1 Crossbreak Active Timer
        [2]   // Ribbon Washer Brush #2 Crossbreak Active Timer
        [6]   // Ribbon Washer Spray #3 Off Timer
   T95 : TIMER[2] := ([0].PRE := 1000, [0].ACC := 790, [0].EN := 1, [0].TT := 1, [1].PRE := 300000, [1].ACC := 279330, [1].EN := 1, [1].TT := 1);
        [0]   // LEHR SPEED Sample period Timer
        [0].DN   // LEHR SPEED Sample Period timer Elapsed
        [1]   // LEHR SPEED Long term Lehr speed Record interval Timer
        [1].DN   // LEHR SPEED Long term Lehr speed Record interval Timer
   TMP_d : DINT := 32767; {access Read Only}
   TMP_dDirection : DINT;
   TMP_dIndex : DINT := 501;
   TMP_dMacIndex : DINT := 20;
   TMP_Index : DINT := 32; {access Read Only}
   TMP_r : REAL;
   TMP_rAcc : REAL := 30000.0;
   TMP_rDec : REAL := 30000.0;
   TMP_rSpeed : REAL := 166.66667;
   TMP_rTarget_M1 : REAL;
   TMP_xAlwaysOFF : BOOL; {access Read Only}
   TMP_xDebugOFF : BOOL; {access Read Only}
   TMP_xRun : BOOL;
   TMP_xTestCycle : BOOL;
   To_Cullet : DINT[10] := ([2] := -28087, [3] := -28096, [4] := -28667, [5] := 16, [6] := -28672); {produced}
   TONY : ALIAS FOR B3[10].15;
   TRIM_2IN_PULSE : ALIAS FOR B73[0].2;
   TRIM_SPEED : ALIAS FOR N60[2];
   VHSC_BTR : ALIAS FOR BT41_000;
   VHSC_BTR_E : ALIAS FOR BT41_000.EN;
   VHSC_BTW : ALIAS FOR BT41_001;
   VHSC_CNFG : ALIAS FOR N42[71].0;
   VHSC_MODEBITS_W : ALIAS FOR N42[3];
   VHSC_OUT00_EN : ALIAS FOR N42[2].0;
   VHSC_OUT00_FRC : ALIAS FOR N42[2].8;
   VHSC_OUT01_EN : ALIAS FOR N42[2].1;
   VHSC_OUT01_FRC : ALIAS FOR N42[2].9;
   VHSC_OUT02_EN : ALIAS FOR N42[2].2;
   VHSC_OUT02_FRC : ALIAS FOR N42[2].10;
   VHSC_OUT03_EN : ALIAS FOR N42[2].3;
   VHSC_OUT03_FRC : ALIAS FOR N42[2].11;
   VHSC_OUT04_EN : ALIAS FOR N42[2].4;
   VHSC_OUT04_FRC : ALIAS FOR N42[2].12;
   VHSC_OUT05_EN : ALIAS FOR N42[2].5;
   VHSC_OUT05_FRC : ALIAS FOR N42[2].13;
   VHSC_OUT06_EN : ALIAS FOR N42[2].6;
   VHSC_OUT06_FRC : ALIAS FOR N42[2].14;
   VHSC_OUT07_EN : ALIAS FOR N42[2].7;
   VHSC_OUT07_FRC : ALIAS FOR N42[2].15;
   VHSC_OUT0_OFLSD : ALIAS FOR N42[29];
   VHSC_OUT0_OFMSD : ALIAS FOR N42[28];
   VHSC_OUT0_ONLSD : ALIAS FOR N42[27];
   VHSC_OUT0_ONMSD : ALIAS FOR N42[26];
   VHSC_OUT1_OFLSD : ALIAS FOR N42[34];
   VHSC_OUT1_OFMSD : ALIAS FOR N42[33];
   VHSC_OUT1_ONLSD : ALIAS FOR N42[32];
   VHSC_OUT1_ONMSD : ALIAS FOR N42[31];
   VHSC_OUT2_OFLSD : ALIAS FOR N42[39];
   VHSC_OUT2_OFMSD : ALIAS FOR N42[38];
   VHSC_OUT2_ONLSD : ALIAS FOR N42[37];
   VHSC_OUT2_ONMSD : ALIAS FOR N42[36];
   VHSC_OUT4_OFLSD : ALIAS FOR N42[49];
   VHSC_OUT4_OFMSD : ALIAS FOR N42[48];
   VHSC_OUT4_ONLSD : ALIAS FOR N42[47];
   VHSC_OUT4_ONMSD : ALIAS FOR N42[46];
   VHSC_OUT6_OFLSD : ALIAS FOR N42[59];
   VHSC_OUT6_OFMSD : ALIAS FOR N42[58];
   VHSC_OUT6_ONLSD : ALIAS FOR N42[57];
   VHSC_OUT6_ONMSD : ALIAS FOR N42[56];
   VHSC_OUT7_OFLSD : ALIAS FOR N42[64];
   VHSC_OUT7_OFMSD : ALIAS FOR N42[63];
   VHSC_OUT7_ONLSD : ALIAS FOR N42[62];
   VHSC_OUT7_ONMSD : ALIAS FOR N42[61];
   VHSC_PC00_LOADP : ALIAS FOR N42[1].8;
   VHSC_PC00_LPRE : ALIAS FOR N42[14];
   VHSC_PC00_LROLL : ALIAS FOR N42[6];
   VHSC_PC00_MPRE : ALIAS FOR N42[13];
   VHSC_PC00_MROLL : ALIAS FOR N42[5];
   VHSC_PC00_PERIO : ALIAS FOR N42[21];
   VHSC_PC01_LOADP : ALIAS FOR N42[1].9;
   VHSC_PC01_LPRE : ALIAS FOR N42[16];
   VHSC_PC01_LROLL : ALIAS FOR N42[8];
   VHSC_PC01_MPRE : ALIAS FOR N42[15];
   VHSC_PC01_MROLL : ALIAS FOR N42[7];
   VHSC_PC01_PERIO : ALIAS FOR N42[22];
   VHSC_PC02_LOADP : ALIAS FOR N42[1].10;
   VHSC_PC02_LPRE : ALIAS FOR N42[18];
   VHSC_PC02_LROLL : ALIAS FOR N42[10];
   VHSC_PC02_MPRE : ALIAS FOR N42[17];
   VHSC_PC02_MROLL : ALIAS FOR N42[9];
   VHSC_PC02_PERIO : ALIAS FOR N42[23];
   VHSC_PC03_LOADP : ALIAS FOR N42[1].11;
   VHSC_PC03_LPRE : ALIAS FOR N42[19];
   VHSC_PC03_LROLL : ALIAS FOR N42[12];
   VHSC_PC03_MROLL : ALIAS FOR N42[11];
   VHSC_PC03_PERIO : ALIAS FOR N42[24];
   VHSC_STAT : ALIAS FOR N42[71];
   VHSC_WR_EN : ALIAS FOR BT41_001.EN;
   VMCC_M1_AMBER : ALIAS FOR O[67].5;
   VMCC_M1_BLUE : ALIAS FOR O[67].4;
   VMCC_M1_RED : ALIAS FOR O[67].3;
   VMCC_W1_AMBER : ALIAS FOR O[47].5;
   VMCC_W1_BLUE : ALIAS FOR O[47].4;
   VMCC_W1_RED : ALIAS FOR O[47].3;
   VMCCMB_ALM_HRN : ALIAS FOR O[20].3;
   VP917060_MED : ALIAS FOR O[116].14;
   VP917060_THICK : ALIAS FOR O[116].15;
   VP917060_THIN : ALIAS FOR O[116].13;
   VP917065_MED : ALIAS FOR O[114].5;
   VP917065_THICK : ALIAS FOR O[114].6;
   VP917065_THIN : ALIAS FOR O[114].4;
   VP917066_MED : ALIAS FOR O[114].2;
   VP917066_THICK : ALIAS FOR O[114].3;
   VP917066_THIN : ALIAS FOR O[114].1;
   VP917067_MED : ALIAS FOR O[113].15;
   VP917067_THICK : ALIAS FOR O[114].0;
   VP917067_THIN : ALIAS FOR O[113].14;
   VP917068_THICK : ALIAS FOR O[116].7;
   VP917069_THICK : ALIAS FOR O[116].2;
   VP917070_MED : ALIAS FOR O[114].8;
   VP917070_MMI : ALIAS FOR N54[376].9;
   VP917070_THICK : ALIAS FOR O[114].9;
   VP917070_THIN : ALIAS FOR O[114].7;
   VP917071_MED : ALIAS FOR O[114].11;
   VP917071_MMI : ALIAS FOR N54[376].8;
   VP917071_THICK : ALIAS FOR O[114].12;
   VP917071_THIN : ALIAS FOR O[114].10;
   VP917072_MED : ALIAS FOR O[116].11;
   VP917072_THICK : ALIAS FOR O[116].12;
   VP917072_THIN : ALIAS FOR O[116].10;
   VP917073_MED : ALIAS FOR O[115].14;
   VP917073_THICK : ALIAS FOR O[115].15;
   VP917073_THIN : ALIAS FOR O[115].13;
   VP917074_MED : ALIAS FOR O[115].11;
   VP917074_THICK : ALIAS FOR O[115].12;
   VP917074_THIN : ALIAS FOR O[115].10;
   VP917075_MED : ALIAS FOR O[115].8;
   VP917075_THICK : ALIAS FOR O[115].9;
   VP917075_THIN : ALIAS FOR O[115].7;
   VP917076_MED : ALIAS FOR O[115].5;
   VP917076_THICK : ALIAS FOR O[115].6;
   VP917076_THIN : ALIAS FOR O[115].4;
   VP917077_MED : ALIAS FOR O[114].14;
   VP917077_THICK : ALIAS FOR O[114].15;
   VP917077_THIN : ALIAS FOR O[114].13;
   W1_ALM_RESET : ALIAS FOR I[42].9;
   W1_ALM_SILENCE : ALIAS FOR I[42].8;
   W1_COMM_PWR : ALIAS FOR I[42].11;
   W1_DC_INPWR : ALIAS FOR I[42].2;
   W1_DC_OUTPWR : ALIAS FOR I[42].3;
   W1_DC_PS1 : ALIAS FOR I[42].6;
   W1_DC_PS2 : ALIAS FOR I[42].7;
   W1_DRV_CONT_ON : ALIAS FOR I[42].1;
   W1_DRV_FLT_LMP : ALIAS FOR O[47].1;
   W1_DRV_FLT_RES : ALIAS FOR O[47].2;
   W1_ESTOP : ALIAS FOR I[42].10;
   W1_ESTOPPWR : ALIAS FOR I[42].5;
   W_APC_ACTIVE : ALIAS FOR W_B3[0].10;
   W_APC_BUTTON : ALIAS FOR W_I[8].10;
   W_APC_FILL_DONE : ALIAS FOR W_T4[20];
   W_B3 : DINT[7] := ([0] := 2#0000_0000_0000_0000_0000_0000_0001_0110, [6] := 2#0000_0000_0000_0000_0000_0000_0001_0000);
        [0].1   // Shutdown Latch Enable/Disable Washer
        [0].10   // APC Tank Fill Cycle Activated
        [0].2   // Run Washer System
        [0].3   // Signal to Start Pump CP2A Motor
        [0].4   // Signal to Start Pump CP2B Motor
        [0].5   // Enable Drives CP1A & CP1B
        [0].6   // Signal to Start Pump CP1A Motor
        [0].7   // Signal to Start Pump CP1B Motor
        [0].8   // PWT_LL_LATCH
        [0].9   // Flow Enabled
        [2].0   // Artificial PI Controller Permissive (No Analog Output)
        [2].1   // Eclipse On Permissive
        [2].2   // Eclipse Off Permissive
        [3].2   // Signal for Spare Pump To Start
        [4].0   // Process Water One Shot to Swith Active Pump
        [4].1   // Process Water RO Pump 1 Tank Low Level Limit Switch ONS
        [4].2   // Process Water RO Pump 1 Allow to Run
        [4].3   // Process Water RO Pump 2 Allow to Run
        [6].4   // RO System Pump Motor Signal to Start
   W_BLOW_PID_TIMER : ALIAS FOR W_T4[15];
   W_BLOWDOWN_ACTIVE : ALIAS FOR W_T4[18];
   W_BLOWDOWN_TIMER : ALIAS FOR W_T4[17];
   W_BLOWDOWN_VALVE : ALIAS FOR W_O[10].12;
   W_C5 : COUNTER[1] := ([0].PRE := 100, [0].ACC := 7359, [0].CU := 1, [0].DN := 1);
        [0]   // Process Water Counter to Switch Active Pump
   W_CB1_AUXILLARY : ALIAS FOR W_I[8].12;
   W_CB1_PID_TIMER : ALIAS FOR W_T4[9];
   W_CB1_START : ALIAS FOR W_O[10].1;
   W_CB2_AUXILLARY : ALIAS FOR W_I[8].11;
   W_CB2_START : ALIAS FOR W_O[10].3;
   W_COMPUTE_TCD3 : ALIAS FOR W_N7[923];
   W_COMPUTE_TCD5B : ALIAS FOR W_N7[926];
   W_CONDUCT_SENSOR : ALIAS FOR W_N7[110];
